// TIA Portal project "proiect" (V17) (continued)
   END_STEP
   TRANSITION Trans117 FROM Step105 TO Step106   // T117
      := "LS.  mixer_spate";
   END_TRANSITION
   STEP Step106:   // S106, max time T#10S, warning time T#7S
              R    "DB_Markers_Auto".step1_left
   END_STEP
   TRANSITION Trans118 FROM Step106 TO Initializare1   // T118, jump
      := NOT "DB_06_Write_Arduino".Stepper1_left AND NOT "DB_HMI_buttons"."Start/Stop_proces_auto";
   END_TRANSITION
   STEP Step107:   // S107, max time T#10S, warning time T#7S
      // stepper up-down
              S    "DB_Markers_Auto".step2_down
   END_STEP
   TRANSITION Trans119 FROM Step107 TO Step108   // T119
      := "LS. mixer_jos";
   END_TRANSITION
   STEP Step108:   // S108, max time T#10S, warning time T#7S
              R    "DB_Markers_Auto".step2_down
   END_STEP
   TRANSITION Trans120 FROM Step108 TO Step124   // T120
      := NOT "DB_06_Write_Arduino".Stepper2_down;
   END_TRANSITION
   STEP Step109:   // S109, max time T#10S, warning time T#7S
      // stepper oriz
              S    "DB_Markers_Auto".step1_left
   END_STEP
   TRANSITION Trans121 FROM Step109 TO Step110   // T121
      := "LS.  mixer_spate";
   END_TRANSITION
   STEP Step110:   // S110, max time T#10S, warning time T#7S
              R    "DB_Markers_Auto".step1_left
   END_STEP
   TRANSITION Trans122 FROM Step110 TO Initializare1   // T122, jump
      := NOT "DB_06_Write_Arduino".Stepper1_left AND NOT "DB_HMI_buttons"."Start/Stop_proces_auto";
   END_TRANSITION
   STEP Step111:   // S111, max time T#10S, warning time T#7S
              S    "DB_Markers_Auto".step2_down
   END_STEP
   TRANSITION Trans123 FROM Step111 TO Step112   // T123
      := "LS. mixer_jos";
   END_TRANSITION
   STEP Step112:   // S112, max time T#10S, warning time T#7S
              R    "DB_Markers_Auto".step2_down
   END_STEP
   TRANSITION Trans124 FROM Step112 TO Step125   // T124
      := NOT "DB_06_Write_Arduino".Stepper2_down;
   END_TRANSITION
   STEP Step113:   // S113, max time T#10S, warning time T#7S
              S    "DB_Markers_Auto".step1_left
   END_STEP
   TRANSITION Trans125 FROM Step113 TO Step114   // T125
      := "LS.  mixer_spate";
   END_TRANSITION
   STEP Step114:   // S114, max time T#10S, warning time T#7S
              R    "DB_Markers_Auto".step1_left
   END_STEP
   TRANSITION Trans126 FROM Step114 TO Initializare1   // T126, jump
      := NOT "DB_06_Write_Arduino".Stepper1_left AND NOT "DB_HMI_buttons"."Start/Stop_proces_auto";
   END_TRANSITION
   STEP Step115:   // S115, max time T#10S, warning time T#7S
              S    "DB_Markers_Auto".step2_down
   END_STEP
   TRANSITION Trans127 FROM Step115 TO Step116   // T127
      := "LS. mixer_jos";
   END_TRANSITION
   STEP Step116:   // S116, max time T#10S, warning time T#7S
              R    "DB_Markers_Auto".step2_down
   END_STEP
   TRANSITION Trans128 FROM Step116 TO Step126   // T128
      := NOT "DB_06_Write_Arduino".Stepper2_down;
   END_TRANSITION
   STEP Step117:   // S117, max time T#10S, warning time T#7S
              S    "DB_Markers_Auto".step1_left
   END_STEP
   TRANSITION Trans129 FROM Step117 TO Step118   // T129
      := "LS.  mixer_spate";
   END_TRANSITION
   STEP Step118:   // S118, max time T#10S, warning time T#7S
              R    "DB_Markers_Auto".step1_left
   END_STEP
   TRANSITION Trans130 FROM Step118 TO Initializare1   // T130, jump
      := NOT "DB_06_Write_Arduino".Stepper1_left AND "DB_HMI_buttons"."Start/Stop_proces_auto";
   END_TRANSITION
   STEP Step121:   // S121, max time T#10S, warning time T#7S
   END_STEP
   TRANSITION Trans135 FROM Step121 TO Initializare1   // T135, jump
      := "DB_HMI"."MAN/AUTO";
   END_TRANSITION
   STEP Step124:   // S124, max time T#10S, warning time T#7S
              D    "delay7",t#5s
   END_STEP
   TRANSITION Trans138 FROM Step124 TO Step42   // T138
      := "delay7";
   END_TRANSITION
   STEP Step123:   // S123, max time T#10S, warning time T#7S
              D    "delay7",t#5s
   END_STEP
   TRANSITION Trans137 FROM Step123 TO "On mixer"   // T137
      := "delay7";
   END_TRANSITION
   STEP Step125:   // S125, max time T#10S, warning time T#7S
              D    "delay7", t#5s
   END_STEP
   TRANSITION Trans139 FROM Step125 TO Step24   // T139
      := "delay7";
   END_TRANSITION
   STEP Step126:   // S126, max time T#10S, warning time T#7S
              D    "delay7",  t#5s
   END_STEP
   TRANSITION Trans140 FROM Step126 TO "On mixer2"   // T140
      := "delay7";
   END_TRANSITION
END_FUNCTION_BLOCK

// folder: FC-uri

FUNCTION "FC_outputs" : Void   // FC1, LAD
TITLE = outputs
{ S7_Optimized_Access := 'TRUE' }
VERSION : 0.1
BEGIN

REGION Network 1: releu plita
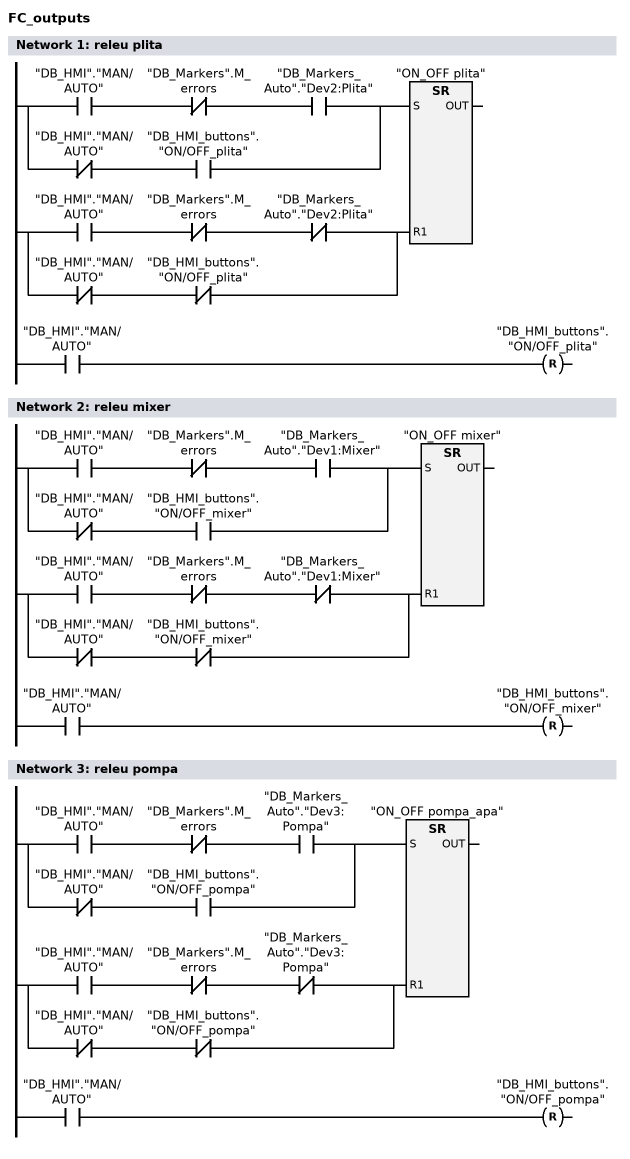
   RUNG wire#powerrail
      Contact( "DB_HMI"."MAN/AUTO" )
      I_Contact( "DB_Markers".M_errors )
      Contact( "DB_Markers_Auto"."Dev2:Plita" )
      wire#w1
      S_SR(operand := "ON_OFF plita", r1 := wire#w2)
   END_RUNG
   RUNG wire#powerrail
      I_Contact( "DB_HMI"."MAN/AUTO" )
      Contact( "DB_HMI_buttons"."ON/OFF_plita" )
   END_RUNG wire#w1
   RUNG wire#powerrail
      Contact( "DB_HMI"."MAN/AUTO" )
      I_Contact( "DB_Markers".M_errors )
      I_Contact( "DB_Markers_Auto"."Dev2:Plita" )
   END_RUNG wire#w2
   RUNG wire#powerrail
      I_Contact( "DB_HMI"."MAN/AUTO" )
      I_Contact( "DB_HMI_buttons"."ON/OFF_plita" )
   END_RUNG wire#w2
   RUNG wire#powerrail
      Contact( "DB_HMI"."MAN/AUTO" )
      R_Coil( "DB_HMI_buttons"."ON/OFF_plita" )
   END_RUNG
   // the same network as SCL:
   IF ("DB_HMI"."MAN/AUTO" AND NOT "DB_Markers".M_errors AND "DB_Markers_Auto"."Dev2:Plita") OR (NOT "DB_HMI"."MAN/AUTO" AND "DB_HMI_buttons"."ON/OFF_plita") THEN
       "ON_OFF plita" := TRUE;   // SR flip-flop
   END_IF;
   IF ("DB_HMI"."MAN/AUTO" AND NOT "DB_Markers".M_errors AND NOT "DB_Markers_Auto"."Dev2:Plita") OR (NOT "DB_HMI"."MAN/AUTO" AND NOT "DB_HMI_buttons"."ON/OFF_plita") THEN
       "ON_OFF plita" := FALSE;
   END_IF;
   IF "DB_HMI"."MAN/AUTO" THEN "DB_HMI_buttons"."ON/OFF_plita" := FALSE; END_IF;
END_REGION

REGION Network 2: releu mixer
   RUNG wire#powerrail
      Contact( "DB_HMI"."MAN/AUTO" )
      I_Contact( "DB_Markers".M_errors )
      Contact( "DB_Markers_Auto"."Dev1:Mixer" )
      wire#w1
      S_SR(operand := "ON_OFF mixer", r1 := wire#w2)
   END_RUNG
   RUNG wire#powerrail
      I_Contact( "DB_HMI"."MAN/AUTO" )
      Contact( "DB_HMI_buttons"."ON/OFF_mixer" )
   END_RUNG wire#w1
   RUNG wire#powerrail
      Contact( "DB_HMI"."MAN/AUTO" )
      I_Contact( "DB_Markers".M_errors )
      I_Contact( "DB_Markers_Auto"."Dev1:Mixer" )
   END_RUNG wire#w2
   RUNG wire#powerrail
      I_Contact( "DB_HMI"."MAN/AUTO" )
      I_Contact( "DB_HMI_buttons"."ON/OFF_mixer" )
   END_RUNG wire#w2
   RUNG wire#powerrail
      Contact( "DB_HMI"."MAN/AUTO" )
      R_Coil( "DB_HMI_buttons"."ON/OFF_mixer" )
   END_RUNG
   // the same network as SCL:
   IF ("DB_HMI"."MAN/AUTO" AND NOT "DB_Markers".M_errors AND "DB_Markers_Auto"."Dev1:Mixer") OR (NOT "DB_HMI"."MAN/AUTO" AND "DB_HMI_buttons"."ON/OFF_mixer") THEN
       "ON_OFF mixer" := TRUE;   // SR flip-flop
   END_IF;
   IF ("DB_HMI"."MAN/AUTO" AND NOT "DB_Markers".M_errors AND NOT "DB_Markers_Auto"."Dev1:Mixer") OR (NOT "DB_HMI"."MAN/AUTO" AND NOT "DB_HMI_buttons"."ON/OFF_mixer") THEN
       "ON_OFF mixer" := FALSE;
   END_IF;
   IF "DB_HMI"."MAN/AUTO" THEN "DB_HMI_buttons"."ON/OFF_mixer" := FALSE; END_IF;
END_REGION

REGION Network 3: releu pompa
   RUNG wire#powerrail
      Contact( "DB_HMI"."MAN/AUTO" )
      I_Contact( "DB_Markers".M_errors )
      Contact( "DB_Markers_Auto"."Dev3:Pompa" )
      wire#w1
      S_SR(operand := "ON_OFF pompa_apa", r1 := wire#w2)
   END_RUNG
   RUNG wire#powerrail
      I_Contact( "DB_HMI"."MAN/AUTO" )
      Contact( "DB_HMI_buttons"."ON/OFF_pompa" )
   END_RUNG wire#w1
   RUNG wire#powerrail
      Contact( "DB_HMI"."MAN/AUTO" )
      I_Contact( "DB_Markers".M_errors )
      I_Contact( "DB_Markers_Auto"."Dev3:Pompa" )
   END_RUNG wire#w2
   RUNG wire#powerrail
      I_Contact( "DB_HMI"."MAN/AUTO" )
      I_Contact( "DB_HMI_buttons"."ON/OFF_pompa" )
   END_RUNG wire#w2
   RUNG wire#powerrail
      Contact( "DB_HMI"."MAN/AUTO" )
      R_Coil( "DB_HMI_buttons"."ON/OFF_pompa" )
   END_RUNG
   // the same network as SCL:
   IF ("DB_HMI"."MAN/AUTO" AND NOT "DB_Markers".M_errors AND "DB_Markers_Auto"."Dev3:Pompa") OR (NOT "DB_HMI"."MAN/AUTO" AND "DB_HMI_buttons"."ON/OFF_pompa") THEN
       "ON_OFF pompa_apa" := TRUE;   // SR flip-flop
   END_IF;
   IF ("DB_HMI"."MAN/AUTO" AND NOT "DB_Markers".M_errors AND NOT "DB_Markers_Auto"."Dev3:Pompa") OR (NOT "DB_HMI"."MAN/AUTO" AND NOT "DB_HMI_buttons"."ON/OFF_pompa") THEN
       "ON_OFF pompa_apa" := FALSE;
   END_IF;
   IF "DB_HMI"."MAN/AUTO" THEN "DB_HMI_buttons"."ON/OFF_pompa" := FALSE; END_IF;
END_REGION
END_FUNCTION

FUNCTION "FC_messages" : Void   // FC2, LAD
TITLE = MESSAGES
{ S7_Optimized_Access := 'TRUE' }
VERSION : 0.1
BEGIN

REGION Network 1: Initializare
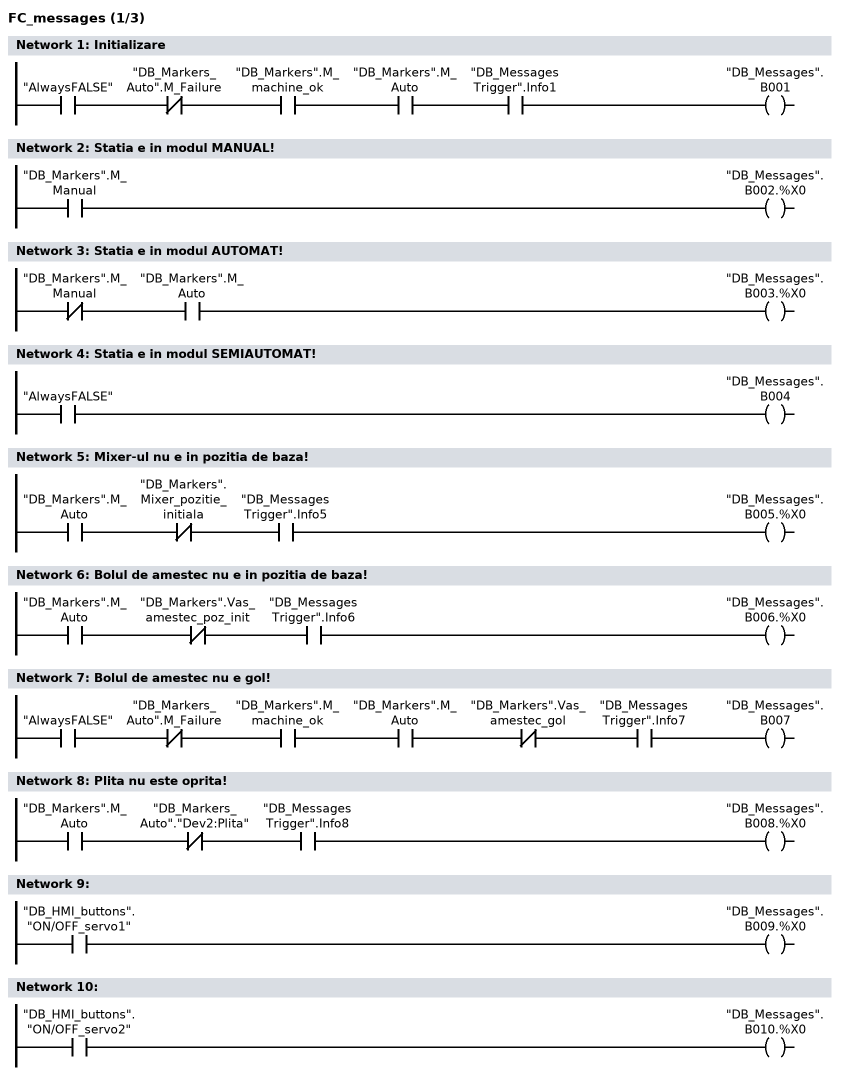
   RUNG wire#powerrail
      Contact( "AlwaysFALSE" )
      I_Contact( "DB_Markers_Auto".M_Failure )
      Contact( "DB_Markers".M_machine_ok )
      Contact( "DB_Markers".M_Auto )
      Contact( "DB_MessagesTrigger".Info1 )
      Coil( "DB_Messages".B001 )
   END_RUNG
   // the same network as SCL:
   "DB_Messages".B001 := "AlwaysFALSE" AND NOT "DB_Markers_Auto".M_Failure AND "DB_Markers".M_machine_ok AND "DB_Markers".M_Auto AND "DB_MessagesTrigger".Info1;
END_REGION

REGION Network 2: Statia e in modul MANUAL!
   RUNG wire#powerrail
      Contact( "DB_Markers".M_Manual )
      Coil( "DB_Messages".B002.%X0 )
   END_RUNG
   // the same network as SCL:
   "DB_Messages".B002.%X0 := "DB_Markers".M_Manual;
END_REGION

REGION Network 3: Statia e in modul AUTOMAT!
   RUNG wire#powerrail
      I_Contact( "DB_Markers".M_Manual )
      Contact( "DB_Markers".M_Auto )
      Coil( "DB_Messages".B003.%X0 )
   END_RUNG
   // the same network as SCL:
   "DB_Messages".B003.%X0 := NOT "DB_Markers".M_Manual AND "DB_Markers".M_Auto;
END_REGION

REGION Network 4: Statia e in modul SEMIAUTOMAT!
   RUNG wire#powerrail
      Contact( "AlwaysFALSE" )
      Coil( "DB_Messages".B004 )
   END_RUNG
   // the same network as SCL:
   "DB_Messages".B004 := "AlwaysFALSE";
END_REGION

REGION Network 5: Mixer-ul nu e in pozitia de baza!
   RUNG wire#powerrail
      Contact( "DB_Markers".M_Auto )
      I_Contact( "DB_Markers".Mixer_pozitie_initiala )
      Contact( "DB_MessagesTrigger".Info5 )
      Coil( "DB_Messages".B005.%X0 )
   END_RUNG
   // the same network as SCL:
   "DB_Messages".B005.%X0 := "DB_Markers".M_Auto AND NOT "DB_Markers".Mixer_pozitie_initiala AND "DB_MessagesTrigger".Info5;
END_REGION

REGION Network 6: Bolul de amestec nu e in pozitia de baza!
   RUNG wire#powerrail
      Contact( "DB_Markers".M_Auto )
      I_Contact( "DB_Markers".Vas_amestec_poz_init )
      Contact( "DB_MessagesTrigger".Info6 )
      Coil( "DB_Messages".B006.%X0 )
   END_RUNG
   // the same network as SCL:
   "DB_Messages".B006.%X0 := "DB_Markers".M_Auto AND NOT "DB_Markers".Vas_amestec_poz_init AND "DB_MessagesTrigger".Info6;
END_REGION

REGION Network 7: Bolul de amestec nu e gol!
   RUNG wire#powerrail
      Contact( "AlwaysFALSE" )
      I_Contact( "DB_Markers_Auto".M_Failure )
      Contact( "DB_Markers".M_machine_ok )
      Contact( "DB_Markers".M_Auto )
      I_Contact( "DB_Markers".Vas_amestec_gol )
      Contact( "DB_MessagesTrigger".Info7 )
      Coil( "DB_Messages".B007 )
   END_RUNG
   // the same network as SCL:
   "DB_Messages".B007 := "AlwaysFALSE" AND NOT "DB_Markers_Auto".M_Failure AND "DB_Markers".M_machine_ok AND "DB_Markers".M_Auto AND NOT "DB_Markers".Vas_amestec_gol AND "DB_MessagesTrigger".Info7;
END_REGION

REGION Network 8: Plita nu este oprita!
   RUNG wire#powerrail
      Contact( "DB_Markers".M_Auto )
      I_Contact( "DB_Markers_Auto"."Dev2:Plita" )
      Contact( "DB_MessagesTrigger".Info8 )
      Coil( "DB_Messages".B008.%X0 )
   END_RUNG
   // the same network as SCL:
   "DB_Messages".B008.%X0 := "DB_Markers".M_Auto AND NOT "DB_Markers_Auto"."Dev2:Plita" AND "DB_MessagesTrigger".Info8;
END_REGION

REGION Network 9
   RUNG wire#powerrail
      Contact( "DB_HMI_buttons"."ON/OFF_servo1" )
      Coil( "DB_Messages".B009.%X0 )
   END_RUNG
   // the same network as SCL:
   "DB_Messages".B009.%X0 := "DB_HMI_buttons"."ON/OFF_servo1";
END_REGION

REGION Network 10
   RUNG wire#powerrail
      Contact( "DB_HMI_buttons"."ON/OFF_servo2" )
      Coil( "DB_Messages".B010.%X0 )
   END_RUNG
   // the same network as SCL:
   "DB_Messages".B010.%X0 := "DB_HMI_buttons"."ON/OFF_servo2";
END_REGION

REGION Network 11: stepper 1 in functionare
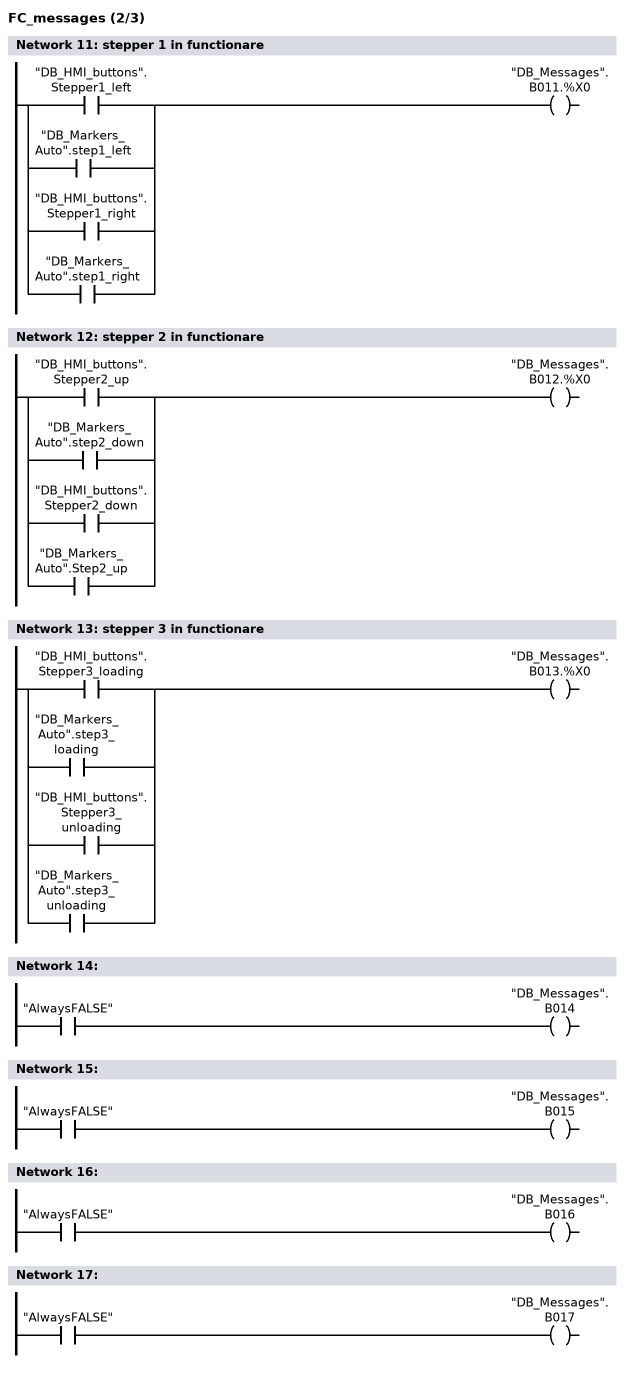
   RUNG wire#powerrail
      Contact( "DB_HMI_buttons".Stepper1_left )
      wire#w1
      Coil( "DB_Messages".B011.%X0 )
   END_RUNG
   RUNG wire#powerrail
      Contact( "DB_Markers_Auto".step1_left )
   END_RUNG wire#w1
   RUNG wire#powerrail
      Contact( "DB_HMI_buttons".Stepper1_right )
   END_RUNG wire#w1
   RUNG wire#powerrail
      Contact( "DB_Markers_Auto".step1_right )
   END_RUNG wire#w1
   // the same network as SCL:
   "DB_Messages".B011.%X0 := "DB_HMI_buttons".Stepper1_left OR "DB_Markers_Auto".step1_left OR "DB_HMI_buttons".Stepper1_right OR "DB_Markers_Auto".step1_right;
END_REGION

REGION Network 12: stepper 2 in functionare
   RUNG wire#powerrail
      Contact( "DB_HMI_buttons".Stepper2_up )
      wire#w1
      Coil( "DB_Messages".B012.%X0 )
   END_RUNG
   RUNG wire#powerrail
      Contact( "DB_Markers_Auto".step2_down )
   END_RUNG wire#w1
   RUNG wire#powerrail
      Contact( "DB_HMI_buttons".Stepper2_down )
   END_RUNG wire#w1
   RUNG wire#powerrail
      Contact( "DB_Markers_Auto".Step2_up )
   END_RUNG wire#w1
   // the same network as SCL:
   "DB_Messages".B012.%X0 := "DB_HMI_buttons".Stepper2_up OR "DB_Markers_Auto".step2_down OR "DB_HMI_buttons".Stepper2_down OR "DB_Markers_Auto".Step2_up;
END_REGION

REGION Network 13: stepper 3 in functionare
   RUNG wire#powerrail
      Contact( "DB_HMI_buttons".Stepper3_loading )
      wire#w1
      Coil( "DB_Messages".B013.%X0 )
   END_RUNG
   RUNG wire#powerrail
      Contact( "DB_Markers_Auto".step3_loading )
   END_RUNG wire#w1
   RUNG wire#powerrail
      Contact( "DB_HMI_buttons".Stepper3_unloading )
   END_RUNG wire#w1
   RUNG wire#powerrail
      Contact( "DB_Markers_Auto".step3_unloading )
   END_RUNG wire#w1
   // the same network as SCL:
   "DB_Messages".B013.%X0 := "DB_HMI_buttons".Stepper3_loading OR "DB_Markers_Auto".step3_loading OR "DB_HMI_buttons".Stepper3_unloading OR "DB_Markers_Auto".step3_unloading;
END_REGION

REGION Network 14
   RUNG wire#powerrail
      Contact( "AlwaysFALSE" )
      Coil( "DB_Messages".B014 )
   END_RUNG
   // the same network as SCL:
   "DB_Messages".B014 := "AlwaysFALSE";
END_REGION

REGION Network 15
   RUNG wire#powerrail
      Contact( "AlwaysFALSE" )
      Coil( "DB_Messages".B015 )
   END_RUNG
   // the same network as SCL:
   "DB_Messages".B015 := "AlwaysFALSE";
END_REGION

REGION Network 16
   RUNG wire#powerrail
      Contact( "AlwaysFALSE" )
      Coil( "DB_Messages".B016 )
   END_RUNG
   // the same network as SCL:
   "DB_Messages".B016 := "AlwaysFALSE";
END_REGION

REGION Network 17
   RUNG wire#powerrail
      Contact( "AlwaysFALSE" )
      Coil( "DB_Messages".B017 )
   END_RUNG
   // the same network as SCL:
   "DB_Messages".B017 := "AlwaysFALSE";
END_REGION

REGION Network 18
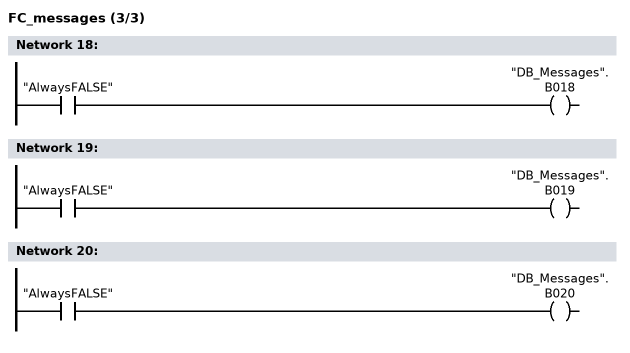
   RUNG wire#powerrail
      Contact( "AlwaysFALSE" )
      Coil( "DB_Messages".B018 )
   END_RUNG
   // the same network as SCL:
   "DB_Messages".B018 := "AlwaysFALSE";
END_REGION

REGION Network 19
   RUNG wire#powerrail
      Contact( "AlwaysFALSE" )
      Coil( "DB_Messages".B019 )
   END_RUNG
   // the same network as SCL:
   "DB_Messages".B019 := "AlwaysFALSE";
END_REGION

REGION Network 20
   RUNG wire#powerrail
      Contact( "AlwaysFALSE" )
      Coil( "DB_Messages".B020 )
   END_RUNG
   // the same network as SCL:
   "DB_Messages".B020 := "AlwaysFALSE";
END_REGION
END_FUNCTION

FUNCTION "FC_Markers" : Void   // FC3, LAD
TITLE = limite/pozitii initiale
{ S7_Optimized_Access := 'TRUE' }
VERSION : 0.1
BEGIN

REGION Network 1: machine ok
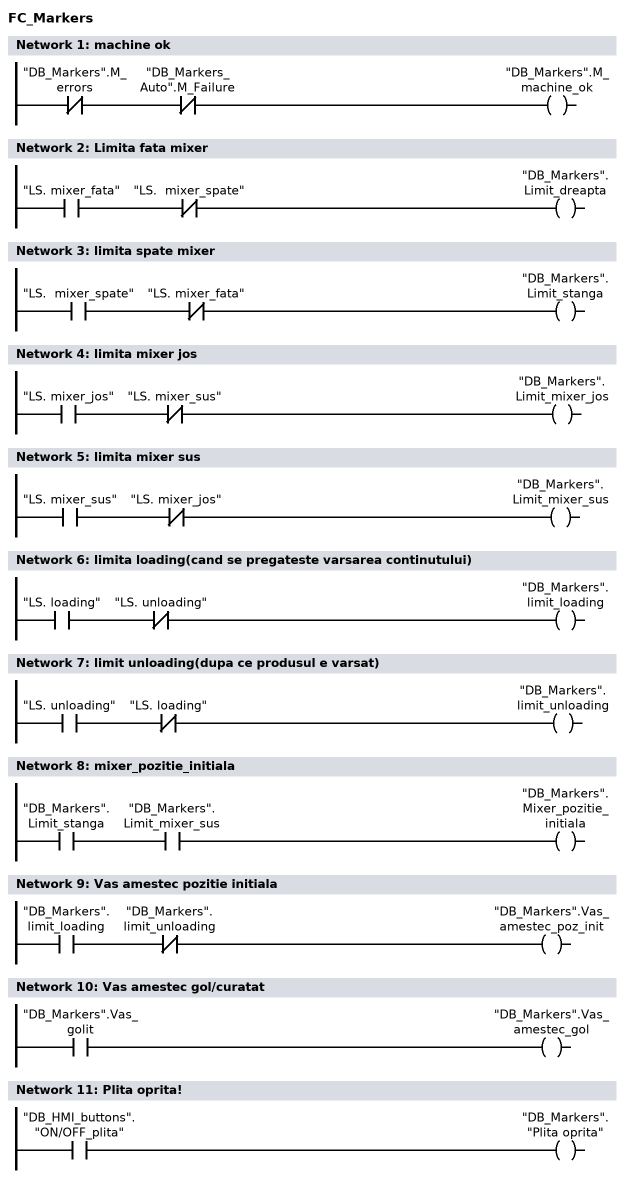
   RUNG wire#powerrail
      I_Contact( "DB_Markers".M_errors )
      I_Contact( "DB_Markers_Auto".M_Failure )
      Coil( "DB_Markers".M_machine_ok )
   END_RUNG
   // the same network as SCL:
   "DB_Markers".M_machine_ok := NOT "DB_Markers".M_errors AND NOT "DB_Markers_Auto".M_Failure;
END_REGION

REGION Network 2: Limita fata mixer
   RUNG wire#powerrail
      Contact( "LS. mixer_fata" )
      I_Contact( "LS.  mixer_spate" )
      Coil( "DB_Markers".Limit_dreapta )
   END_RUNG
   // the same network as SCL:
   "DB_Markers".Limit_dreapta := "LS. mixer_fata" AND NOT "LS.  mixer_spate";
END_REGION

REGION Network 3: limita spate mixer
   RUNG wire#powerrail
      Contact( "LS.  mixer_spate" )
      I_Contact( "LS. mixer_fata" )
      Coil( "DB_Markers".Limit_stanga )
   END_RUNG
   // the same network as SCL:
   "DB_Markers".Limit_stanga := "LS.  mixer_spate" AND NOT "LS. mixer_fata";
END_REGION

REGION Network 4: limita mixer jos
   RUNG wire#powerrail
      Contact( "LS. mixer_jos" )
      I_Contact( "LS. mixer_sus" )
      Coil( "DB_Markers".Limit_mixer_jos )
   END_RUNG
   // the same network as SCL:
   "DB_Markers".Limit_mixer_jos := "LS. mixer_jos" AND NOT "LS. mixer_sus";
END_REGION

REGION Network 5: limita mixer sus
   RUNG wire#powerrail
      Contact( "LS. mixer_sus" )
      I_Contact( "LS. mixer_jos" )
      Coil( "DB_Markers".Limit_mixer_sus )
   END_RUNG
   // the same network as SCL:
   "DB_Markers".Limit_mixer_sus := "LS. mixer_sus" AND NOT "LS. mixer_jos";
END_REGION

REGION Network 6: limita loading(cand se pregateste varsarea continutului)
   RUNG wire#powerrail
      Contact( "LS. loading" )
      I_Contact( "LS. unloading" )
      Coil( "DB_Markers".limit_loading )
   END_RUNG
   // the same network as SCL:
   "DB_Markers".limit_loading := "LS. loading" AND NOT "LS. unloading";
END_REGION

REGION Network 7: limit unloading(dupa ce produsul e varsat)
   RUNG wire#powerrail
      Contact( "LS. unloading" )
      I_Contact( "LS. loading" )
      Coil( "DB_Markers".limit_unloading )
   END_RUNG
   // the same network as SCL:
   "DB_Markers".limit_unloading := "LS. unloading" AND NOT "LS. loading";
END_REGION

REGION Network 8: mixer_pozitie_initiala
   RUNG wire#powerrail
      Contact( "DB_Markers".Limit_stanga )
      Contact( "DB_Markers".Limit_mixer_sus )
      Coil( "DB_Markers".Mixer_pozitie_initiala )
   END_RUNG
   // the same network as SCL:
   "DB_Markers".Mixer_pozitie_initiala := "DB_Markers".Limit_stanga AND "DB_Markers".Limit_mixer_sus;
END_REGION

REGION Network 9: Vas amestec pozitie initiala
   RUNG wire#powerrail
      Contact( "DB_Markers".limit_loading )
      I_Contact( "DB_Markers".limit_unloading )
      Coil( "DB_Markers".Vas_amestec_poz_init )
   END_RUNG
   // the same network as SCL:
   "DB_Markers".Vas_amestec_poz_init := "DB_Markers".limit_loading AND NOT "DB_Markers".limit_unloading;
END_REGION

REGION Network 10: Vas amestec gol/curatat
   RUNG wire#powerrail
      Contact( "DB_Markers".Vas_golit )
      Coil( "DB_Markers".Vas_amestec_gol )
   END_RUNG
   // the same network as SCL:
   "DB_Markers".Vas_amestec_gol := "DB_Markers".Vas_golit;
END_REGION

REGION Network 11: Plita oprita!
   RUNG wire#powerrail
      Contact( "DB_HMI_buttons"."ON/OFF_plita" )
      Coil( "DB_Markers"."Plita oprita" )
   END_RUNG
   // the same network as SCL:
   "DB_Markers"."Plita oprita" := "DB_HMI_buttons"."ON/OFF_plita";
END_REGION
END_FUNCTION

FUNCTION "FC_Errors" : Void   // FC4, LAD
TITLE = ERORI
{ S7_Optimized_Access := 'TRUE' }
VERSION : 0.1
BEGIN

REGION Network 1 (SCL): Error marker/Failure marker
   IF  "DB_Errors"."Eroare1:Vas in aer" AND "DB_Errors"."Eroare2:Mixer" AND "DB_Errors"."Eroare3:temp plita" AND "DB_Errors"."Eroare4:Servo oprite" THEN
       // Statement section IF
       "DB_Markers".M_errors := TRUE;
       "DB_Markers_Auto".M_Failure:=TRUE
       ;
   END_IF;
END_REGION

REGION Network 2: STOP : ciuperca activata
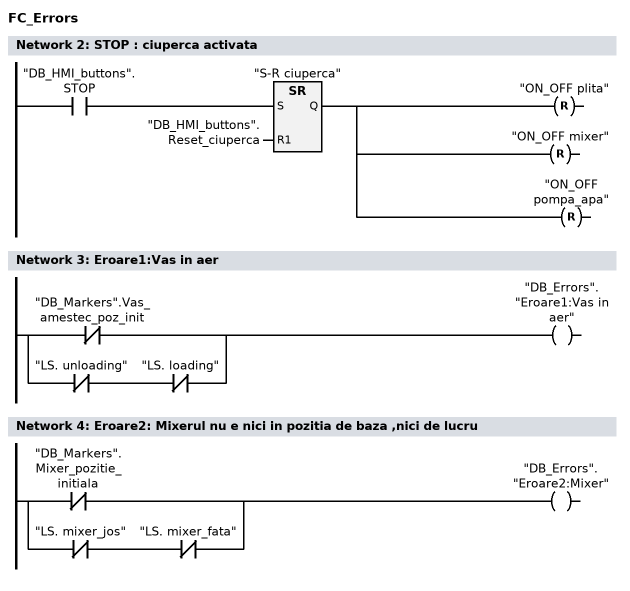
   RUNG wire#powerrail
      Contact( "DB_HMI_buttons".STOP )
      S_SR(operand := "S-R ciuperca", r1 := "DB_HMI_buttons".Reset_ciuperca)
      wire#w1
      R_Coil( "ON_OFF plita" )
   END_RUNG
   RUNG wire#w1
      R_Coil( "ON_OFF mixer" )
   END_RUNG
   RUNG wire#w1
      R_Coil( "ON_OFF pompa_apa" )
   END_RUNG
   // the same network as SCL:
   IF "DB_HMI_buttons".STOP THEN
       "S-R ciuperca" := TRUE;   // SR flip-flop
   END_IF;
   IF "DB_HMI_buttons".Reset_ciuperca THEN "S-R ciuperca" := FALSE; END_IF;
   IF "S-R ciuperca" THEN
       "ON_OFF plita" := FALSE;
       "ON_OFF mixer" := FALSE;
       "ON_OFF pompa_apa" := FALSE;
   END_IF;
END_REGION

REGION Network 3: Eroare1:Vas in aer
   RUNG wire#powerrail
      I_Contact( "DB_Markers".Vas_amestec_poz_init )
      wire#w1
      Coil( "DB_Errors"."Eroare1:Vas in aer" )
   END_RUNG
   RUNG wire#powerrail
      I_Contact( "LS. unloading" )
      I_Contact( "LS. loading" )
   END_RUNG wire#w1
   // the same network as SCL:
   "DB_Errors"."Eroare1:Vas in aer" := NOT "DB_Markers".Vas_amestec_poz_init OR (NOT "LS. unloading" AND NOT "LS. loading");
END_REGION

REGION Network 4: Eroare2: Mixerul nu e nici in pozitia de baza ,nici de lucru
   RUNG wire#powerrail
      I_Contact( "DB_Markers".Mixer_pozitie_initiala )
      wire#w1
      Coil( "DB_Errors"."Eroare2:Mixer" )
   END_RUNG
   RUNG wire#powerrail
      I_Contact( "LS. mixer_jos" )
      I_Contact( "LS. mixer_fata" )
   END_RUNG wire#w1
   // the same network as SCL:
   "DB_Errors"."Eroare2:Mixer" := NOT "DB_Markers".Mixer_pozitie_initiala OR (NOT "LS. mixer_jos" AND NOT "LS. mixer_fata");
END_REGION
END_FUNCTION

FUNCTION "FC_Mod_manual" : Void   // FC6, LAD
TITLE = M0D_MANUAL
{ S7_Optimized_Access := 'TRUE' }
VERSION : 0.1
   VAR_TEMP   // added for the SCL form of the ladder/FBD networks
      _w1 : Bool;
      _w2 : Bool;
   END_VAR
BEGIN

REGION Network 1: setare bit 1 pentru SERVO1
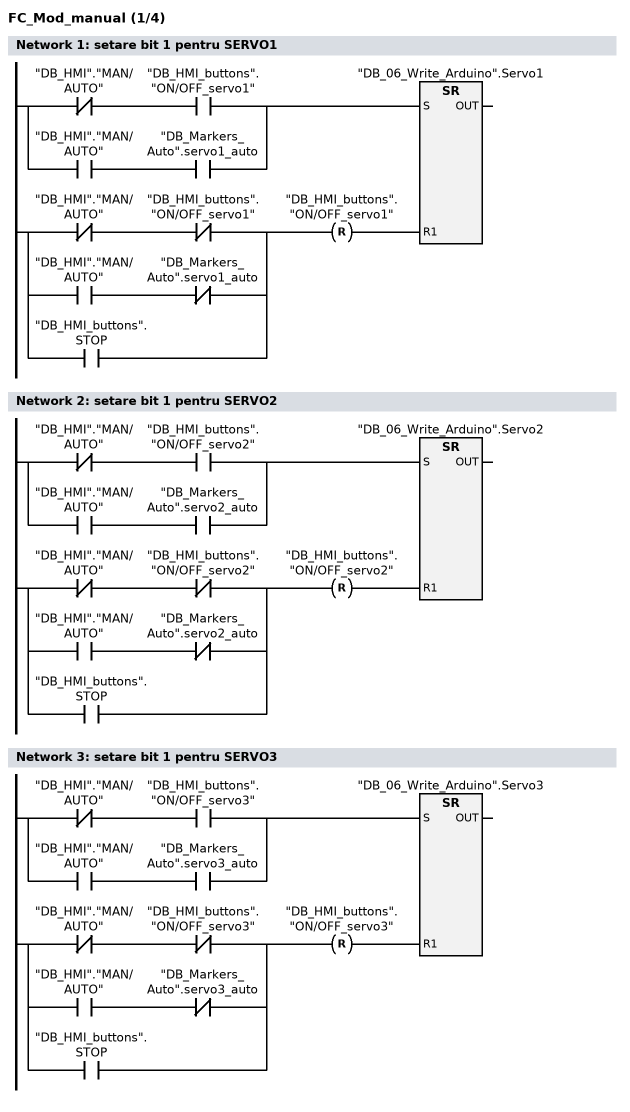
   RUNG wire#powerrail
      I_Contact( "DB_HMI"."MAN/AUTO" )
      Contact( "DB_HMI_buttons"."ON/OFF_servo1" )
      wire#w1
      S_SR(operand := "DB_06_Write_Arduino".Servo1, r1 := wire#w3)
   END_RUNG
   RUNG wire#powerrail
      Contact( "DB_HMI"."MAN/AUTO" )
      Contact( "DB_Markers_Auto".servo1_auto )
   END_RUNG wire#w1
   RUNG wire#powerrail
      I_Contact( "DB_HMI"."MAN/AUTO" )
      I_Contact( "DB_HMI_buttons"."ON/OFF_servo1" )
      wire#w2
      R_Coil( "DB_HMI_buttons"."ON/OFF_servo1" )
   END_RUNG wire#w3
   RUNG wire#powerrail
      Contact( "DB_HMI"."MAN/AUTO" )
      I_Contact( "DB_Markers_Auto".servo1_auto )
   END_RUNG wire#w2
   RUNG wire#powerrail
      Contact( "DB_HMI_buttons".STOP )
   END_RUNG wire#w2
   // the same network as SCL:
   #_w1 := (NOT "DB_HMI"."MAN/AUTO" AND NOT "DB_HMI_buttons"."ON/OFF_servo1") OR ("DB_HMI"."MAN/AUTO" AND NOT "DB_Markers_Auto".servo1_auto) OR "DB_HMI_buttons".STOP;
   #_w2 := (NOT "DB_HMI"."MAN/AUTO" AND "DB_HMI_buttons"."ON/OFF_servo1") OR ("DB_HMI"."MAN/AUTO" AND "DB_Markers_Auto".servo1_auto);
   IF #_w1 THEN "DB_HMI_buttons"."ON/OFF_servo1" := FALSE; END_IF;
   IF #_w2 THEN
       "DB_06_Write_Arduino".Servo1 := TRUE;   // SR flip-flop
   END_IF;
   IF #_w1 THEN "DB_06_Write_Arduino".Servo1 := FALSE; END_IF;
END_REGION

REGION Network 2: setare bit 1 pentru SERVO2
   RUNG wire#powerrail
      I_Contact( "DB_HMI"."MAN/AUTO" )
      Contact( "DB_HMI_buttons"."ON/OFF_servo2" )
      wire#w1
      S_SR(operand := "DB_06_Write_Arduino".Servo2, r1 := wire#w3)
   END_RUNG
   RUNG wire#powerrail
      Contact( "DB_HMI"."MAN/AUTO" )
      Contact( "DB_Markers_Auto".servo2_auto )
   END_RUNG wire#w1
   RUNG wire#powerrail
      I_Contact( "DB_HMI"."MAN/AUTO" )
      I_Contact( "DB_HMI_buttons"."ON/OFF_servo2" )
      wire#w2
      R_Coil( "DB_HMI_buttons"."ON/OFF_servo2" )
   END_RUNG wire#w3
   RUNG wire#powerrail
      Contact( "DB_HMI"."MAN/AUTO" )
      I_Contact( "DB_Markers_Auto".servo2_auto )
   END_RUNG wire#w2
   RUNG wire#powerrail
      Contact( "DB_HMI_buttons".STOP )
   END_RUNG wire#w2
   // the same network as SCL:
   #_w1 := (NOT "DB_HMI"."MAN/AUTO" AND NOT "DB_HMI_buttons"."ON/OFF_servo2") OR ("DB_HMI"."MAN/AUTO" AND NOT "DB_Markers_Auto".servo2_auto) OR "DB_HMI_buttons".STOP;
   #_w2 := (NOT "DB_HMI"."MAN/AUTO" AND "DB_HMI_buttons"."ON/OFF_servo2") OR ("DB_HMI"."MAN/AUTO" AND "DB_Markers_Auto".servo2_auto);
   IF #_w1 THEN "DB_HMI_buttons"."ON/OFF_servo2" := FALSE; END_IF;
   IF #_w2 THEN
       "DB_06_Write_Arduino".Servo2 := TRUE;   // SR flip-flop
   END_IF;
   IF #_w1 THEN "DB_06_Write_Arduino".Servo2 := FALSE; END_IF;
END_REGION

REGION Network 3: setare bit 1 pentru SERVO3
   RUNG wire#powerrail
      I_Contact( "DB_HMI"."MAN/AUTO" )
      Contact( "DB_HMI_buttons"."ON/OFF_servo3" )
      wire#w1
      S_SR(operand := "DB_06_Write_Arduino".Servo3, r1 := wire#w3)
   END_RUNG
   RUNG wire#powerrail
      Contact( "DB_HMI"."MAN/AUTO" )
      Contact( "DB_Markers_Auto".servo3_auto )
   END_RUNG wire#w1
   RUNG wire#powerrail
      I_Contact( "DB_HMI"."MAN/AUTO" )
      I_Contact( "DB_HMI_buttons"."ON/OFF_servo3" )
      wire#w2
      R_Coil( "DB_HMI_buttons"."ON/OFF_servo3" )
   END_RUNG wire#w3
   RUNG wire#powerrail
      Contact( "DB_HMI"."MAN/AUTO" )
      I_Contact( "DB_Markers_Auto".servo3_auto )
   END_RUNG wire#w2
   RUNG wire#powerrail
      Contact( "DB_HMI_buttons".STOP )
   END_RUNG wire#w2
   // the same network as SCL:
   #_w1 := (NOT "DB_HMI"."MAN/AUTO" AND NOT "DB_HMI_buttons"."ON/OFF_servo3") OR ("DB_HMI"."MAN/AUTO" AND NOT "DB_Markers_Auto".servo3_auto) OR "DB_HMI_buttons".STOP;
   #_w2 := (NOT "DB_HMI"."MAN/AUTO" AND "DB_HMI_buttons"."ON/OFF_servo3") OR ("DB_HMI"."MAN/AUTO" AND "DB_Markers_Auto".servo3_auto);
   IF #_w1 THEN "DB_HMI_buttons"."ON/OFF_servo3" := FALSE; END_IF;
   IF #_w2 THEN
       "DB_06_Write_Arduino".Servo3 := TRUE;   // SR flip-flop
   END_IF;
   IF #_w1 THEN "DB_06_Write_Arduino".Servo3 := FALSE; END_IF;
END_REGION

REGION Network 4: setare bit 1 pentru SERVO4
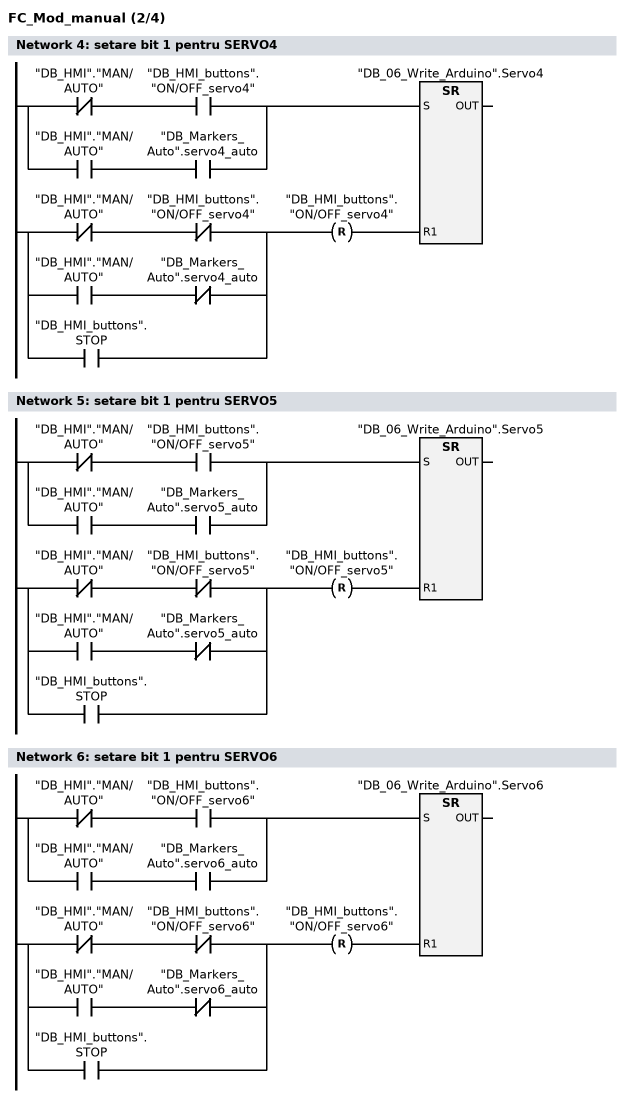
   RUNG wire#powerrail
      I_Contact( "DB_HMI"."MAN/AUTO" )
      Contact( "DB_HMI_buttons"."ON/OFF_servo4" )
      wire#w1
      S_SR(operand := "DB_06_Write_Arduino".Servo4, r1 := wire#w3)
   END_RUNG
   RUNG wire#powerrail
      Contact( "DB_HMI"."MAN/AUTO" )
      Contact( "DB_Markers_Auto".servo4_auto )
   END_RUNG wire#w1
   RUNG wire#powerrail
      I_Contact( "DB_HMI"."MAN/AUTO" )
      I_Contact( "DB_HMI_buttons"."ON/OFF_servo4" )
      wire#w2
      R_Coil( "DB_HMI_buttons"."ON/OFF_servo4" )
   END_RUNG wire#w3
   RUNG wire#powerrail
      Contact( "DB_HMI"."MAN/AUTO" )
      I_Contact( "DB_Markers_Auto".servo4_auto )
   END_RUNG wire#w2
   RUNG wire#powerrail
      Contact( "DB_HMI_buttons".STOP )
   END_RUNG wire#w2
   // the same network as SCL:
   #_w1 := (NOT "DB_HMI"."MAN/AUTO" AND NOT "DB_HMI_buttons"."ON/OFF_servo4") OR ("DB_HMI"."MAN/AUTO" AND NOT "DB_Markers_Auto".servo4_auto) OR "DB_HMI_buttons".STOP;
   #_w2 := (NOT "DB_HMI"."MAN/AUTO" AND "DB_HMI_buttons"."ON/OFF_servo4") OR ("DB_HMI"."MAN/AUTO" AND "DB_Markers_Auto".servo4_auto);
   IF #_w1 THEN "DB_HMI_buttons"."ON/OFF_servo4" := FALSE; END_IF;
   IF #_w2 THEN
       "DB_06_Write_Arduino".Servo4 := TRUE;   // SR flip-flop
   END_IF;
   IF #_w1 THEN "DB_06_Write_Arduino".Servo4 := FALSE; END_IF;
END_REGION

REGION Network 5: setare bit 1 pentru SERVO5
   RUNG wire#powerrail
      I_Contact( "DB_HMI"."MAN/AUTO" )
      Contact( "DB_HMI_buttons"."ON/OFF_servo5" )
      wire#w1
      S_SR(operand := "DB_06_Write_Arduino".Servo5, r1 := wire#w3)
   END_RUNG
   RUNG wire#powerrail
      Contact( "DB_HMI"."MAN/AUTO" )
      Contact( "DB_Markers_Auto".servo5_auto )
   END_RUNG wire#w1
   RUNG wire#powerrail
      I_Contact( "DB_HMI"."MAN/AUTO" )
      I_Contact( "DB_HMI_buttons"."ON/OFF_servo5" )
      wire#w2
      R_Coil( "DB_HMI_buttons"."ON/OFF_servo5" )
   END_RUNG wire#w3
   RUNG wire#powerrail
      Contact( "DB_HMI"."MAN/AUTO" )
      I_Contact( "DB_Markers_Auto".servo5_auto )
   END_RUNG wire#w2
   RUNG wire#powerrail
      Contact( "DB_HMI_buttons".STOP )
   END_RUNG wire#w2
   // the same network as SCL:
   #_w1 := (NOT "DB_HMI"."MAN/AUTO" AND NOT "DB_HMI_buttons"."ON/OFF_servo5") OR ("DB_HMI"."MAN/AUTO" AND NOT "DB_Markers_Auto".servo5_auto) OR "DB_HMI_buttons".STOP;
   #_w2 := (NOT "DB_HMI"."MAN/AUTO" AND "DB_HMI_buttons"."ON/OFF_servo5") OR ("DB_HMI"."MAN/AUTO" AND "DB_Markers_Auto".servo5_auto);
   IF #_w1 THEN "DB_HMI_buttons"."ON/OFF_servo5" := FALSE; END_IF;
   IF #_w2 THEN
       "DB_06_Write_Arduino".Servo5 := TRUE;   // SR flip-flop
   END_IF;
   IF #_w1 THEN "DB_06_Write_Arduino".Servo5 := FALSE; END_IF;
END_REGION

